   	   
   	    If Not IsDate(restore_time) Then
   			bfde4b54-0db7-4817-8032-87127bf19bb9 "Can't set f(x) view time to <" & restore_time & ">."
   		End If
   		
   		'---------------------------------------------------------
   		            
   	    ' go through the whole file, copy line by line, and replace the two archive variable names:
   	    While Not f2.eof
   			restore_entry=f2.lineinputstring
   			restore_entry= Replace(restore_entry, source_name1, target_name1)
   			restore_entry= Replace(restore_entry, source_name2, target_name2)
   			restore_entry= Replace(restore_entry, source_name3, target_name3)
   			restore_entry= Replace(restore_entry, source_name4, target_name4)
   			restore_entry= Replace(restore_entry, source_name5, target_name5)
   			restore_entry= Replace(restore_entry, source_name6, target_name6)
   			restore_entry= Replace(restore_entry, source_name7, target_name7)
   			restore_entry= Replace(restore_entry, source_name8, target_name8)
   			restore_entry= Replace(restore_entry, source_name9, target_name9)
   			f.lineprint(restore_entry)		
   		Wend
   		
   		f2.Close
   	    f.Close
   	       
   	    bb0abc73-aec8-40d0-9880-0280a6a3de42
   		Delay(2)
   		bec8f1e5-2ab1-45f6-ad91-1d37c469eb91 0502_Trend Historical, 0
   	            
   	    bfde4b54-0db7-4817-8032-87127bf19bb9 "Restored archive <" & archive_path & "> to <" & current_path &"> at " & restore_time & "."
   	    
   	    Set f2= Nothing
   	    Set f= Nothing
   		Else
   			
   		bb0abc73-aec8-40d0-9880-0280a6a3de42
   		bfde4b54-0db7-4817-8032-87127bf19bb9 "Long-term archive <" & archive_path & "> not found."
   	End If
   	
       Set fs= Nothing
       

VB script "LHmiView_vbsFECreateFolder"
   On Error Resume Next
   
   '-----------------------DEFINE PARAMETERS-------------------------------------------
   'kindOfOperatingSystem: 0 = Windows, 1 = Windows CE
   ' tempFs: Reference on temporary fileSystem Object
   ' fs: Reference on fileSystem Object
   ' f: Reference on file Object
   Dim kindOfOperatingSystem, tempFs, f, fs, file
   
   '--------------------Prove which Operating System is running------------------------
   'Set tempFs = CreateObject("Scripting.FileSystemObject")
   
   'If Err.Number = 0 Then
   '	kindOfOperatingSystem = 0 'Windows / PC based
   'Else
   	kindOfOperatingSystem = 1 'Windows CE / Panel based
   'End If
   
   Set tempFs= Nothing
   Err.Clear
   
   '-----------------create new folder-----------------------
   Dim newfolder
   
   If SmartTags("NewFolder") = "" Then 
     SmartTags("FEStatus") = "Folder name empty"
     Exit Sub
   End If
   
   newfolder = SmartTags("Folder") & SmartTags("NewFolder")
   
   'Windows CE / Panel based
   If kindOfOperatingSystem Then    
     Set fs = CreateObject("FileCtl.FileSystem")
     If fs.Dir(newfolder) = "" Then
       fs.MkDir(newfolder)
       If Err.Number = 0 Then
         SmartTags("FEStatus") = "Folder " & newfolder & " created"
       Else
         SmartTags("FEStatus") = "Could not create folder " & newfolder
       End If
     Else
       SmartTags("FEStatus") = "Folder exists already"
     End If
     
   ' Windows / PC based
   Else
     Set fs = CreateObject("Scripting.FileSystemObject")
     If fs.FolderExists(newfolder) = False Then
       fs.CreateFolder(newfolder)
       If Err.Number = 0 Then
         SmartTags("FEStatus") = "Folder " & newfolder & " created"
       Else
         SmartTags("FEStatus") = "Could not create folder " & newfolder
       End If
     Else
       SmartTags("FEStatus") = "Folder exists already"
     End If
   End If
   
   Set fs = Nothing
   
   LHmiView_vbsFEReadFilesOfFolder SmartTags("Folder")
   LHmiView_vbsFEWriteFilePropertiesToTags SmartTags("index")

VB script "LHmiView_vbsFEDelete"
   On Error Resume Next
   
   '-----------------------DEFINE PARAMETERS-------------------------------------------
   'kindOfOperatingSystem: 0 = Windows, 1 = Windows CE
   ' tempFs: Reference on temporary fileSystem Object
   ' fs: Reference on fileSystem Object
   ' f: Reference on file Object
   Dim kindOfOperatingSystem, tempFs, f, fs, file
   
   '--------------------Prove which Operating System is running------------------------
   'Set tempFs = CreateObject("Scripting.FileSystemObject")
   
   'If Err.Number = 0 Then
   '	kindOfOperatingSystem = 0 'Windows / PC based
   'Else
   	kindOfOperatingSystem = 1 'Windows CE / Panel based
   'End If
   
   Set tempFs= Nothing
   Err.Clear
   
   '-------------------------------Delete folder/file---------------------------------
   Dim i
   
   SmartTags("FEStatus") = "Deleting file..."
   i = SmartTags("fileChosen")
   
   ' Windows CE / Panel based
   If kindOfOperatingSystem Then    
     Set fs = CreateObject("FileCtl.FileSystem")
     Set f = CreateObject("FileCtl.File")
     If i > 0 And SmartTags("File_"&i) <> "" Then
       If SmartTags("isFolder_"&i) <> 0 Then
         fs.RmDir SmartTags("File_"&i)
         If Err.Number = 0 Then
           SmartTags("FEStatus") = "File / Folder deleted: " & SmartTags("File_"&i) 
           SmartTags("File_"&i) = ""
         Else
           SmartTags("FEStatus") = "Could not delete file / folder: " & SmartTags("File_"&i)
         End If
       Else
         fs.kill SmartTags("File_"&i)
         If Err.Number = 0 Then
           SmartTags("FEStatus") = "File / Folder deleted: " & SmartTags("File_"&i) 
         Else
           SmartTags("FEStatus") = "Could not delete file / folder: " & SmartTags("File_"&i)
         End If
         SmartTags("File_"&i) = ""
       End If
     Else
       SmartTags("FEStatus") = "Choose file / folder"
     End If
     
   ' Windows / PC based
   Else
     Set fs = CreateObject("Scripting.FileSystemObject")
      If i > 0 And SmartTags("File_"&i) <> "" Then
       If SmartTags("isFolder_"&i) <> "False" Then
         fs.DeleteFolder(SmartTags("File_"&i))
         If Err.Number = 0 Then
           SmartTags("FEStatus") = "File / folder deleted: " & SmartTags("File_"&i) 
           SmartTags("File_"&i) = ""
         Else
           SmartTags("FEStatus") = "Could not delete file / folder: " & SmartTags("File_"&i)
         End If
       Else
         fs.DeleteFile(SmartTags("File_"&i))
         If Err.Number = 0 Then
           SmartTags("FEStatus") = "Folder / folder deleted: " & SmartTags("File_"&i) 
         Else
           SmartTags("FEStatus") = "Could not delete file/ folder: " & SmartTags("File_"&i)
         End If
         SmartTags("File_"&i) = ""
       End If
     Else
       SmartTags("FEStatus") = "Choose file / folder"
     End If
   End If
   
   Set fs = Nothing
   Set f = Nothing
   
   LHmiView_vbsFEReadFilesOfFolder SmartTags("Folder")
   LHmiView_vbsFEWriteFilePropertiesToTags SmartTags("index")

VB script "LHmiView_vbsFEMove"
   On Error Resume Next
   
   '-----------------------DEFINE PARAMETERS-------------------------------------------
   'kindOfOperatingSystem: 0 = Windows, 1 = Windows CE
   ' tempFs: Reference on temporary fileSystem Object
   ' fs: Reference on fileSystem Object
   ' f: Reference on file Object
   Dim kindOfOperatingSystem, tempFs, f, fs, file
   
   '--------------------Prove which Operating System is running------------------------
   'Set tempFs = CreateObject("Scripting.FileSystemObject")
   
   'If Err.Number = 0 Then
   '	kindOfOperatingSystem = 0 'Windows / PC based
   'Else
   	kindOfOperatingSystem = 1 'Windows CE / Panel based
   'End If
   
   Set tempFs= Nothing
   Err.Clear
   
   '-------------------------------Move folder/file---------------------------------
   Dim  newpath, singleFile, data
   
   ' Windows CE / Panel based
   If kindOfOperatingSystem Then
     If sender = 1 Then 'button "copy" pressed
   	  If SmartTags("copyusb") = True Then
   		    If SmartTags("aIsFolder_"&SmartTags("AfileChosen")) = 0 Then
   		      SmartTags("bufferFile") = SmartTags("AFile_"&SmartTags("AfileChosen"))
   		      SmartTags("bufferFolder") = SmartTags("AFolder")
   		      SmartTags("bufferCopyCut") = True
   		      SmartTags("bufferIsFolder") = SmartTags("AisFolder_"&SmartTags("AfileChosen"))
   		      SmartTags("FEStatus") = "File " & SmartTags("bufferFile") & " copied"
   		    Else
   		      SmartTags("FEStatus") = "Cannot copy folder"
   			End If
   	  Else
   		   If SmartTags("IsFolder_"&SmartTags("fileChosen")) = 0 Then
   		      SmartTags("bufferFile") = SmartTags("File_"&SmartTags("fileChosen"))
   		      SmartTags("bufferFolder") = SmartTags("Folder")
   		      SmartTags("bufferCopyCut") = True
   		      SmartTags("bufferIsFolder") = SmartTags("isFolder_"&SmartTags("fileChosen"))
   		      SmartTags("FEStatus") = "File " & SmartTags("bufferFile") & " copied"
   		    Else
   		      SmartTags("FEStatus") = "Cannot copy folder"
   		   End If
   	  End If
   	  
     
     ElseIf sender = 3 Then 'button "cut" is pressed
   	  If SmartTags("copyusb") = True Then
   		    SmartTags("bufferFile") = SmartTags("AFile_"&SmartTags("AfileChosen"))
   		    SmartTags("bufferFolder") = SmartTags("AFolder")
   		    SmartTags("bufferCopyCut") = False 
   		    SmartTags("bufferIsFolder") = SmartTags("AisFolder_"&SmartTags("AfileChosen"))
   		    SmartTags("FEStatus") = "File " & SmartTags("bufferFile") & " cut"
   	  Else
   		  	SmartTags("bufferFile") = SmartTags("File_"&SmartTags("fileChosen"))
   		    SmartTags("bufferFolder") = SmartTags("Folder")
   		    SmartTags("bufferCopyCut") = False 
   		    SmartTags("bufferIsFolder") = SmartTags("isFolder_"&SmartTags("fileChosen"))
   		    SmartTags("FEStatus") = "File " & SmartTags("bufferFile") & " cut"   
   	  End If
   	  
   	  
     ElseIf sender = 2 Then 'button "move" pressed
       singleFile = Replace (SmartTags("bufferFile"),  SmartTags("bufferFolder"), "")
       newpath = SmartTags("Folder") & singleFile  
       If SmartTags("bufferCopyCut") = False Then   
         If SmartTags("bufferIsFolder") <> 0 Then
           Set fs = CreateObject("FileCtl.FileSystem")
           fs.MoveFile SmartTags("bufferFile"), newpath
         Else
           Set fs = CreateObject("FileCtl.FileSystem")
           fs.FileCopy SmartTags("bufferFile"), newpath
           fs.kill SmartTags("bufferFile")
         End If
       Else
         Set fs = CreateObject("FileCtl.FileSystem")
         fs.FileCopy SmartTags("bufferFile"), newpath
       End If 
       SmartTags("FEStatus") = "File " & SmartTags("bufferFile") & " pasted"
       LHmiView_vbsFEReadFilesOfFolder SmartTags("Folder")
       LHmiView_vbsFEWriteFilePropertiesToTags SmartTags("index")
     End If
   ' Windows / PC based
   Else
     If sender = 1 Then 'button "copy" pressed
   	  If SmartTags("copyusb") = True Then
   	    SmartTags("bufferFile") = SmartTags("aFile_"&SmartTags("AfileChosen"))
   	    SmartTags("bufferFolder") = SmartTags("AFolder")
   	    SmartTags("bufferCopyCut") = True
   	    SmartTags("bufferIsFolder") = SmartTags("aisFolder_"&SmartTags("AfileChosen"))
   	    SmartTags("FEStatus") = "File " & SmartTags("bufferFile") & " copied"
   	  Else
   		SmartTags("bufferFile") = SmartTags("File_"&SmartTags("fileChosen"))
   	    SmartTags("bufferFolder") = SmartTags("Folder")
   	    SmartTags("bufferCopyCut") = True
   	    SmartTags("bufferIsFolder") = SmartTags("isFolder_"&SmartTags("fileChosen"))
   	    SmartTags("FEStatus") = "File " & SmartTags("bufferFile") & " copied"
   	  End If
   	  
     
     ElseIf sender = 3 Then 'button "cut" is pressed
   	  If SmartTags("copyusb") = True Then
   		    SmartTags("bufferFile") = SmartTags("File_"&SmartTags("AfileChosen"))
   		    SmartTags("bufferFolder") = SmartTags("AFolder")
   		    SmartTags("bufferCopyCut") = False 
   		    SmartTags("bufferIsFolder") = SmartTags("aisFolder_"&SmartTags("AfileChosen"))
   		    SmartTags("FEStatus") = "File " & SmartTags("bufferFile") & " cut"
   	  Else
   		    SmartTags("bufferFile") = SmartTags("File_"&SmartTags("AfileChosen"))
   		    SmartTags("bufferFolder") = SmartTags("AFolder")
   		    SmartTags("bufferCopyCut") = False 
   		    SmartTags("bufferIsFolder") = SmartTags("aisFolder_"&SmartTags("AfileChosen"))
   		    SmartTags("FEStatus") = "File " & SmartTags("bufferFile") & " cut"
   	  End If    
   	  
     ElseIf sender = 2 Then 'button "move" pressed
       singleFile = Replace (SmartTags("bufferFile"),  SmartTags("bufferFolder"), "")
       newpath = SmartTags("Folder") & singleFile  
       Set fs = CreateObject("Scripting.FileSystemObject")
       If SmartTags("bufferCopyCut") = False Then
         If SmartTags("bufferIsFolder") = "True" Then
           data = fs.GetFolder(SmartTags("bufferFile"))
           fs.MoveFolder data, newpath
         Else
           data = fs.GetFile(SmartTags("bufferFile"))
           fs.MoveFile data, newpath
         End If
       Else
         If SmartTags("bufferIsFolder") = "True" Then
           data = fs.GetFolder(SmartTags("bufferFile"))
           fs.CopyFolder data, newpath
         Else
           data = fs.GetFile(SmartTags("bufferFile"))
           fs.CopyFile data, newpath
         End If
       End If
       If Err.Number <> 0 Then
         SmartTags("FEStatus") = Err.Description & "Could not paste file / folder"
       Else
         SmartTags("FEStatus") = "File / Folder " & SmartTags("bufferFile") & " pasted"
       End If
       LHmiView_vbsFEReadFilesOfFolder SmartTags("Folder")
       LHmiView_vbsFEWriteFilePropertiesToTags SmartTags("index")
     End If
   End If

VB script "LHmiView_vbsFEPreviousFolder"
   On Error Resume Next
   
   Dim folder, prevFolder
   
   If SmartTags("Search") = True Then
     SmartTags("Search") = False
     LHmiView_vbsFEReadFilesOfFolder(SmartTags("FEsearchFolder"))
     LHmiView_vbsFEWriteFilePropertiesToTags 1
   Else
   	If Len(SmartTags("Folder")) > 1 Then
   	    folder = Left (SmartTags("Folder"),  InStrRev (SmartTags("Folder"), "\")-1)
   	    prevFolder = Left (folder, InStrRev (folder, "\"))
   	    LHmiView_vbsFEReadFilesOfFolder(prevFolder)
   	    LHmiView_vbsFEWriteFilePropertiesToTags 1
   	    SmartTags("index") = 1
   	    SmartTags("FEStatus") = "Folder " & prevFolder & " opened"
   	Else
   	    SmartTags("FEStatus") = "Operation not possible"
   	End If
   End If

VB script "LHmiView_vbsFEReadFilesOfFolder"
   On Error Resume Next
   
   '-----------------------DEFINE PARAMETERS-------------------------------------------
   'kindOfOperatingSystem: 0 = Windows, 1 = Windows CE
   ' tempFs: Reference on temporary fileSystem Object
   ' fs: Reference on fileSystem Object
   ' f: Reference on file Object
   Dim kindOfOperatingSystem, tempFs, f, fs, file
   
   '--------------------Prove which Operating System is running------------------------
   'Set tempFs = CreateObject("Scripting.FileSystemObject")
   
   'If Err.Number = 0 Then
   '	kindOfOperatingSystem = 0 'Windows / PC based
   'Else
   	kindOfOperatingSystem = 1 'Windows CE / Panel based
   'End If
   
   Set tempFs= Nothing
   Err.Clear
   
   '-------------------------------Read files of folder---------------------------------
   Dim isFolder, counter, index, textStream, folder, dataInFolder, fileList
   
   index = 1
   
   ' Windows CE / Panel based
   If kindOfOperatingSystem Then 
     If folderpar = "" Then
       folderpar = "\"
     End If
        
     Set fs = CreateObject("FileCtl.FileSystem")
     Set f = CreateObject("FileCtl.File")
     If fs.Dir("\flash\106226404_Tools") = "" Then   fs.MkDir("\flash\106226404_Tools")
     f.open "\flash\106226404_Tools\LHmiView_FileList.txt", 2 'textfile where the files are stored
     
     file = fs.dir(folderpar & "*")
     counter = 0
     index = 1
     f.lineprint(folderpar)
     f.lineprint("-1")
     f.LinePrint "#106226404_FE_Site_"&index
     
     Do While file <> "" 
       If (counter < 10) Then  'write 10 files (pathname and isFolder) to textfile
         If ((fs.GetAttr(folderpar & file) And 16) <> 0 ) Then
           isFolder = True
         Else
           isFolder = False
         End If
         f.LinePrint(folderpar & file)
         f.LinePrint(isFolder)
         file = fs.dir
         counter = counter + 1
       Else
         counter = 0
         index = index + 1
         f.LinePrint "#106226404_FE_Site_"&index 
       End If
     Loop
     
     f.Close
     
   ' Windows / PC based
   Else
     If (folderpar = "") Then
       folderpar = "C:\"
     End If
     
     Set fs = CreateObject("Scripting.FileSystemObject")
     fileList = "C:\106226404_Tools\LHmiView_FileList.txt"
     If Not fs.FolderExists("C:\106226404_Tools") Then fs.CreateFolder "C:\106226404_Tools"
     If Not fs.FileExists(fileList) Then fs.CreateTextFile fileList
     Set f = fs.GetFile(fileList)
     Set textStream = f.OpenAsTextStream(2,-2)
     
     counter = 0
     index = 1
     textStream.WriteLine(folderpar)
     textStream.WriteLine("-1")
     textStream.WriteLine "#106226404_FE_Site_"&index
     
     Set folder = fs.GetFolder(folderpar)
     
     Set dataInFolder = folder.SubFolders
     For Each file In dataInFolder
       If Not file.Attributes And 2 Then
         If (counter < 10) Then 'write 10 files (pathname and isFolder) to textfile
           textStream.WriteLine(file.Path)
           textStream.WriteLine("True")
           counter = counter + 1
         Else
           counter = 0
           index = index + 1
           textStream.WriteLine "#106226404_FE_Site_"&index 
         End If
       End If
     Next
     
     Set dataInFolder = folder.Files
     For Each file In dataInFolder
       If Not file.Attributes And 2 Then
         If (counter < 10) Then 'write 10 folder (pathname and isFolder) to textfile
           textStream.WriteLine(file.Path)
           textStream.WriteLine("False")
           counter = counter + 1
         Else
           counter = 0
           index = index + 1
           textStream.WriteLine "#106226404_FE_Site_"&index 
         End If
       End If
     Next
   
     textStream.Close
     Set folder = Nothing
     Set dataInFolder = Nothing
     Set textStream = Nothing
   
   End If
   Set fs = Nothing
   Set f = Nothing

VB script "LHmiView_vbsFERename"
   On Error Resume Next
   
   '-----------------------DEFINE PARAMETERS-------------------------------------------
   'kindOfOperatingSystem: 0 = Windows, 1 = Windows CE
   ' tempFs: Reference on temporary fileSystem Object
   ' fs: Reference on fileSystem Object
   ' f: Reference on file Object
   Dim kindOfOperatingSystem, tempFs, f, fs,file
   
   '--------------------Prove which Operating System is running------------------------
   'Set tempFs = CreateObject("Scripting.FileSystemObject")
   
   'If Err.Number = 0 Then
   '	kindOfOperatingSystem = 0 'Windows / PC based
   'Else
   	kindOfOperatingSystem = 1 'Windows CE / Panel based
   'End If
   
   Set tempFs= Nothing
   Err.Clear
   
   '-------------------------------Rename folder/file---------------------------------
   Dim i, newName, ext, fileName, folder
   
   i = SmartTags("fileChosen")
   fileName = SmartTags("File_"&i)
   
   If fileName <> "" And SmartTags("NewName") <> "" Then
     
     ' Windows CE / Panel based
     If kindOfOperatingSystem Then    
       Set fs = CreateObject("FileCtl.FileSystem")
       If SmartTags("IsFolder_"&i) <> 0 Then 'Rename folder
         newName = SmartTags("Folder") & SmartTags("NewName")
         fs.MoveFile fileName, newName
         If Err.Number = 0 Then
           SmartTags("FEStatus") = "Folder renamed in: " & newName
         Else
           SmartTags("FEStatus") = "Could not rename folder: " & fileName
         End If
       Else 'Keep file extension
         ext = Right(fileName, Len(fileName)-InStrRev(fileName, "."))
         newName = SmartTags("Folder") & SmartTags("NewName") & "." & ext
         fs.MoveFile fileName, newName
         If Err.Number = 0 Then
           SmartTags("FEStatus") = "File renamed in: " & newName
         Else
           SmartTags("FEStatus") = "Could not rename file:" & fileName
         End If    
       End If
       
     ' Windows / PC based
     Else
       Set fs = CreateObject("Scripting.FileSystemObject")
       If SmartTags("IsFolder_"&i) <> "False" Then 'Rename folder
         Set folder = fs.GetFolder(fileName)
         newName = SmartTags("Folder") & SmartTags("NewName")
         fs.MoveFolder fileName, newName
         If Err.Number = 0 Then
           SmartTags("FEStatus") = "Folder renamed in: " & newName
         Else
           SmartTags("FEStatus") = "Error :" & Err.Description & " Could not rename folder: " & fileName
         End If
         Set folder = Nothing
       Else 'Keep file extension
        Set file = fs.GetFile(fileName)
         ext = Right(fileName, Len(fileName)-InStrRev(fileName, "."))
         newName = SmartTags("NewName") & "." & ext
         file.Name = newName
         If Err.Number = 0 Then
           SmartTags("FEStatus") = "File renamed in: " & newName
         Else
           SmartTags("FEStatus") = "Could not rename file: " & fileName
         End If    
         Set file = Nothing
       End If 
     End If
     Set fs = Nothing
    
   Else
     SmartTags("FEStatus") = "No file / folder chosen or name empty"
   End If
   Set fs = Nothing
   LHmiView_vbsFEReadFilesOfFolder SmartTags("Folder")
   LHmiView_vbsFEWriteFilePropertiesToTags SmartTags("index")
     

VB script "LHmiView_vbsFESearch"
   On Error Resume Next
   
   '-----------------------DEFINE PARAMETERS-------------------------------------------
   'kindOfOperatingSystem: 0 = Windows, 1 = Windows CE
   ' tempFs: Reference on temporary fileSystem Object
   ' fs: Reference on fileSystem Object
   ' f: Reference on file Object
   Dim kindOfOperatingSystem, tempFs, f, fs, file
   
   '--------------------Prove which Operating System is running------------------------
   'Set tempFs = CreateObject("Scripting.FileSystemObject")
   
   'If Err.Number = 0 Then
   '	kindOfOperatingSystem = 0 'Windows / PC based
   'Else
   	kindOfOperatingSystem = 1 'Windows CE / Panel based
   'End If
   
   Set tempFs= Nothing
   Err.Clear
   
   '-------------------------------Search folder/file---------------------------------
   Dim i, j, index, line, buffer(), searchString
   
   If SmartTags("FEsearchString") <> "" Then
     SmartTags("FEStatus") = "Searching for text: " & SmartTags("FEsearchString") & "..."
     
     'Windows CE / Panel based
     If kindOfOperatingSystem Then
       Set f = CreateObject("filectl.file")
       Set fs = CreateObject("filectl.Filesystem")
       file = "\flash\106226404_Tools\LHmiView_FileList.txt"
       f.open file, 1 
       i=1
       j=1
       searchString = LCase(SmartTags("FEsearchString")) 
       Do While f.EOF = False 'Check number of lines for Array Definition
         f.LineInputString
         i=i+1
       Loop
       ReDim buffer(i)
       'Reinitialize
       i=1
       f.close
       f.open file,1
       Do While f.EOF = False
         line = LCase(f.LineInputString)
          If InStr(1,line,searchString,0) <> 0 Then
            buffer(i) = line
            buffer(i+1) = f.LineInputString
            i = i+2
            bfde4b54-0db7-4817-8032-87127bf19bb9("Found: "&line)
          End If
       Loop
       f.Close
       If i>1 Then
         SmartTags("FEsearchFolder") = SmartTags("Folder")
         f.open "\flash\106226404_Tools\LHmiView_SearchList.txt", 2  
         index = 1
         f.LinePrint SmartTags("Folder")
         f.LinePrint "#106226404_FE_Site_"&index
         For j=1 To i
           f.LinePrint(buffer(j))
           bfde4b54-0db7-4817-8032-87127bf19bb9("Written: " &buffer(j))
           If (j Mod 20) = 0 Then
             index = index+1
             f.LinePrint "#106226404_FE_Site_"&index
           End If
         Next
         f.close
         fs.kill "\flash\106226404_Tools\LHmiView_FileList.txt"
         fs.FileCopy "\flash\106226404_Tools\LHmiView_SearchList.txt", "\flash\106226404_Tools\LHmiView_FileList.txt"
         fs.kill "\flash\106226404_Tools\LHmiView_SearchList.txt"
         LHmiView_vbsFEWriteFilePropertiesToTags 1
       End If
       SmartTags("FEStatus") = (i-1)/2 & " Files found with text: " & SmartTags("FEsearchString") 
       Set f = Nothing
       Set fs = Nothing
       
     'Windows / PC based
     Else
       Set fs = CreateObject("Scripting.FileSystemObject")
       file = "C:\106226404_Tools\LHmiView_FileList.txt"
       Set f = fs.OpenTextFile (file, 1) 
       i=1
       j=1
       searchString = LCase(SmartTags("FEsearchString")) 
       Do While f.AtEndOfStream <> True 'Check number of lines for Array Definition
         f.ReadLine
         i=i+1
       Loop
       ReDim buffer(i)
       'Reinitialize
       i=1
       f.Close
       Set f = fs.OpenTextFile (file, 1)
       Do While f.AtEndOfStream <> True
         line = LCase(f.ReadLine)
         If InStr(1,line,searchString,0) <> 0 Then
           buffer(i) = line
           buffer(i+1) = f.ReadLine
           i = i+2
         End If
       Loop
       f.Close
       If i>1 Then
         SmartTags("FEsearchFolder") = SmartTags("Folder")
         file = "C:\106226404_Tools\LHmiView_SearchList.txt"
         If Not fs.FileExists(file) Then fs.CreateTextFile file
         Set f = fs.OpenTextFile (file, 2)
         index = 1
         f.WriteLine SmartTags("Folder")
         f.WriteLine "#106226404_FE_Site_"&index
         For j=1 To i
           f.WriteLine(buffer(j))
           bfde4b54-0db7-4817-8032-87127bf19bb9("Written: " &buffer(j))
           If (j Mod 20) = 0 Then
             index = index+1
             f.WriteLine "#106226404_FE_Site_"&index
           End If
         Next
         f.Close
         fs.DeleteFile "C:\106226404_Tools\LHmiView_FileList.txt"
         fs.CopyFile "C:\106226404_Tools\LHmiView_SearchList.txt", "C:\106226404_Tools\LHmiView_FileList.txt"
         fs.DeleteFile "C:\106226404_Tools\LHmiView_SearchList.txt"
         LHmiView_vbsFEWriteFilePropertiesToTags 1
       End If
       SmartTags("FEStatus") = (i-1)/2 & " Files found with text: " & SmartTags("FEsearchString") 
       Set f = Nothing
       Set fs = Nothing          
     End If        
   Else
     SmartTags("FEStatus") = "Search text empty"
   End If      

VB script "LHmiView_vbsFEShowFiles"
   On Error Resume Next
   
   '-----------------------DEFINE PARAMETERS-------------------------------------------
   'kindOfOperatingSystem: 0 = Windows, 1 = Windows CE
   ' tempFs: Reference on temporary fileSystem Object
   ' fs: Reference on fileSystem Object
   ' f: Reference on file Object
   Dim kindOfOperatingSystem, tempFs, f, fs, file
   
   '--------------------Prove which Operating System is running------------------------
   'Set tempFs = CreateObject("Scripting.FileSystemObject")
   
   'If Err.Number = 0 Then
   '	kindOfOperatingSystem = 0 'Windows / PC based
   'Else
   	kindOfOperatingSystem = 1 'Windows CE / Panel based
   'End If
   
   Set tempFs= Nothing
   Err.Clear
   
   '-----------------show files -----------------------
   Dim fileName, ext, obj
   'Windows CE / Panel based
   
   If kindOfOperatingSystem Then  
     If SmartTags("File_"&SmartTags("fileChosen")) <> "" Then
       If SmartTags("IsFolder_"&SmartTags("fileChosen")) <> 0 Then
           LHmiView_vbsFEReadFilesOfFolder(SmartTags("File_"&SmartTags("fileChosen"))&"\")
           LHmiView_vbsFEWriteFilePropertiesToTags 1
           SmartTags("index") = 1
       Else
         fileName = SmartTags("File_"&SmartTags("fileChosen")) 
         ext = LCase(Right(fileName, Len(fileName)-InStrRev(fileName, "."))) 
         fileName = Chr(34) & fileName & Chr(34) ' Add " for spaces in fileName
       ' ExcelViewer: *.xlsx, *.xls, *.xlt
       ' WordViewer: *.docx, *.rtf, *.doc
       ' PdfViewer *.pdf
       ' Internet Explorer *.html
       ' Mediaplayer *.mpa, *.mp2, *.mp3, *.wma, *wav, *.mpg, *.mpeg, *.mpe, *.asf, *.wmv, *.avi
         If ext = "xlsx" Or ext = "xls" Or ext = "xlt" Or _
         ext = "docx" Or ext = "rtf" Or ext = "doc" Or _
         ext = "pdf" Or _
         ext = "html" Or _
         ext = "mpa" Or ext = "mp2" Or ext = "mp3" Or ext = "wma" Or ext = "wav" Or ext = "mpg" Or ext = "mpeg" Or ext = "mpe" Or ext = "asf" Or ext = "wmv" Or ext = "avi" Then
             bf5b406f-e168-4434-a306-9566226aa38b fileName, "", $3$hmiShowNormal$, $3$hmiNo$
         Else
           SmartTags("FEStatus") = "Cannot open file"
         End If  
       End If
     End If
   'Windows / PC based 
   Else
     If SmartTags("File_"&SmartTags("fileChosen")) <> "" Then
       If SmartTags("IsFolder_"&SmartTags("fileChosen")) <> "False" Then
         LHmiView_vbsFEReadFilesOfFolder(SmartTags("File_"&SmartTags("fileChosen"))&"\")
         LHmiView_vbsFEWriteFilePropertiesToTags 1
         SmartTags("index") = 1
       Else  
         fileName = SmartTags("File_"&SmartTags("fileChosen")) 
         Set obj = CreateObject("Wscript.Shell")
         obj.Run fileName
       End If
     Else
       SmartTags("FEStatus") = "No file or folder chosen"
     End If
   End If

VB script "LHmiView_vbsFEWriteFilePropertiesToTags"
   On Error Resume Next
   
   '-----------------------DEFINE PARAMETERS-------------------------------------------
   'kindOfOperatingSystem: 0 = Windows, 1 = Windows CE
   ' tempFs: Reference on temporary fileSystem Object
   ' fs: Reference on fileSystem Object
   ' f: Reference on file Object
   Dim kindOfOperatingSystem, tempFs, f, fs, file
   
   '--------------------Prove which Operating System is running------------------------
   'Set tempFs = CreateObject("Scripting.FileSystemObject")
   
   'If Err.Number = 0 Then
   '	kindOfOperatingSystem = 0 'Windows / PC based
   'Else
   	kindOfOperatingSystem = 1 'Windows CE / Panel based
   'End If
   
   Set tempFs= Nothing
   Err.Clear
   
   '-----------------create new folder-----------------------
   Dim i
   
   If kindOfOperatingSystem Then    
     Set fs = CreateObject("FileCtl.FileSystem")
     Set f = CreateObject("FileCtl.File")
     file = "\flash\106226404_Tools\LHmiView_FileList.txt"
     SmartTags("NextPossible") = True
     If fs.Dir(file) <> "" Then
       f.open file, 1
       SmartTags("Folder") = f.LineInputString
       Do While f.LineInputString <>  "#106226404_FE_Site_"&index  'find current position in file 
       Loop
       
       For i=1 To 10
         If f.EOF = False Then       
           SmartTags("File_" &i) = f.LineInputString
         Else  ' fill tags at the end of the file
           SmartTags("File_" &i) = ""
         End If
         If f.EOF = False Then
           SmartTags("isFolder_" &i) = f.LineInputString
         Else  
           SmartTags("isFolder_" &i) = ""     
         End If
       Next
       
       If f.EOF = True Then
         SmartTags("NextPossible") = False
       Else 
         SmartTags("NextPossible") = True
       End If
       f.Close 
       f.Close
     End If
   ' Windows / PC based
   Else
     Set fs = CreateObject("Scripting.FileSystemObject")
     file = "C:\106226404_Tools\LHmiView_FileList.txt"
     If Not fs.FileExists(file) Then Exit Sub
     Set f = fs.OpenTextFile (file, 1)
     SmartTags("Folder") = f.ReadLine
     Do While f.ReadLine <>  "#106226404_FE_Site_"&index  'find current position in file 
     Loop
     
     For i=1 To 10
       If f.AtEndOfStream = False Then       
         SmartTags("File_" &i) = f.ReadLine
       Else  ' fill tags at the end of the file
         SmartTags("File_" &i) = ""
       End If
       If f.AtEndOfStream = False Then
         SmartTags("isFolder_" &i) = f.ReadLine
       Else  
         SmartTags("isFolder_" &i) = ""     
       End If
     Next
     
     If f.AtEndOfStream = True Then
       SmartTags("NextPossible") = False
     Else 
       SmartTags("NextPossible") = True
     End If
     f.Close    
   End If
   Set fs = Nothing
   Set f = Nothing

VB script "LHmiView_vbsFESearch_1"
   On Error Resume Next
   
   '-----------------------DEFINE PARAMETERS-------------------------------------------
   'kindOfOperatingSystem: 0 = Windows, 1 = Windows CE
   ' tempFs: Reference on temporary fileSystem Object
   ' fs: Reference on fileSystem Object
   ' f: Reference on file Object
   Dim kindOfOperatingSystem, tempFs, f, fs, file
   
   '--------------------Prove which Operating System is running------------------------
   'Set tempFs = CreateObject("Scripting.FileSystemObject")
   
   'If Err.Number = 0 Then
   '	kindOfOperatingSystem = 0 'Windows / PC based
   'Else
   	kindOfOperatingSystem = 1 'Windows CE / Panel based
   'End If
   
   Set tempFs= Nothing
   Err.Clear
   
   '-------------------------------Search folder/file---------------------------------
   Dim i, j, index, line, buffer(), searchString
   
   If SmartTags("AFEsearchString") <> "" Then
     SmartTags("AFEStatus") = "Searching for text: " & SmartTags("AFEsearchString") & "..."
     
     'Windows CE / Panel based
     If kindOfOperatingSystem Then
       Set f = CreateObject("filectl.file")
       Set fs = CreateObject("filectl.Filesystem")
       file = "\flash\106226404_Tools\LHmiView_FileListB.txt"
       f.open file, 1 
       i=1
       j=1
       searchString = LCase(SmartTags("AFEsearchString")) 
       Do While f.EOF = False 'Check number of lines for Array Definition
         f.LineInputString
         i=i+1
       Loop
       ReDim buffer(i)
       'Reinitialize
       i=1
       f.close
       f.open file,1
       Do While f.EOF = False
         line = LCase(f.LineInputString)
          If InStr(1,line,searchString,0) <> 0 Then
            buffer(i) = line
            buffer(i+1) = f.LineInputString
            i = i+2
            bfde4b54-0db7-4817-8032-87127bf19bb9("Found: "&line)
          End If
       Loop
       f.Close
       If i>1 Then
         SmartTags("AFEsearchFolder") = SmartTags("AFolder")
         f.open "\flash\106226404_Tools\LHmiView_SearchListB.txt", 2  
         index = 1
         f.LinePrint SmartTags("AFolder")
         f.LinePrint "#106226404_FE_Site_"&index
         For j=1 To i
           f.LinePrint(buffer(j))
           bfde4b54-0db7-4817-8032-87127bf19bb9("Written: " &buffer(j))
           If (j Mod 20) = 0 Then
             index = index+1
             f.LinePrint "#106226404_FE_Site_"&index
           End If
         Next
         f.close
         fs.kill "\flash\106226404_Tools\LHmiView_FileListB.txt"
         fs.FileCopy "\flash\106226404_Tools\LHmiView_SearchListB.txt", "\flash\106226404_Tools\LHmiView_FileListB.txt"
         fs.kill "\flash\106226404_Tools\LHmiView_SearchListB.txt"
         LHmiView_vbsFEWriteFilePropertiesToTags_1 1
       End If
       SmartTags("AFEStatus") = (i-1)/2 & " Files found with text: " & SmartTags("AFEsearchString") 
       Set f = Nothing
       Set fs = Nothing
       
     'Windows / PC based
     Else
       Set fs = CreateObject("Scripting.FileSystemObject")
       file = "C:\106226404_Tools\LHmiView_FileListB.txt"
       Set f = fs.OpenTextFile (file, 1) 
       i=1
       j=1
       searchString = LCase(SmartTags("AFEsearchString")) 
       Do While f.AtEndOfStream <> True 'Check number of lines for Array Definition
         f.ReadLine
         i=i+1
       Loop
       ReDim buffer(i)
       'Reinitialize
       i=1
       f.Close
       Set f = fs.OpenTextFile (file, 1)
       Do While f.AtEndOfStream <> True
         line = LCase(f.ReadLine)
         If InStr(1,line,searchString,0) <> 0 Then
           buffer(i) = line
           buffer(i+1) = f.ReadLine
           i = i+2
         End If
       Loop
       f.Close
       If i>1 Then
         SmartTags("AFEsearchFolder") = SmartTags("AFolder")
         file = "C:\106226404_Tools\LHmiView_SearchListB.txt"
         If Not fs.FileExists(file) Then fs.CreateTextFile file
         Set f = fs.OpenTextFile (file, 2)
         index = 1
         f.WriteLine SmartTags("AFolder")
         f.WriteLine "#106226404_FE_Site_"&index
         For j=1 To i
           f.WriteLine(buffer(j))
           bfde4b54-0db7-4817-8032-87127bf19bb9("Written: " &buffer(j))
           If (j Mod 20) = 0 Then
             index = index+1
             f.WriteLine "#106226404_FE_Site_"&index
           End If
         Next
         f.Close
         fs.DeleteFile "C:\106226404_Tools\LHmiView_FileListB.txt"
         fs.CopyFile "C:\106226404_Tools\LHmiView_SearchListB.txt", "C:\106226404_Tools\LHmiView_FileListB.txt"
         fs.DeleteFile "C:\106226404_Tools\LHmiView_SearchListB.txt"
         LHmiView_vbsFEWriteFilePropertiesToTags_1 1
       End If
       SmartTags("AFEStatus") = (i-1)/2 & " Files found with text: " & SmartTags("AFEsearchString") 
       Set f = Nothing
       Set fs = Nothing          
     End If        
   Else
     SmartTags("AFEStatus") = "Search text empty"
   End If      

VB script "LHmiView_vbsFEWriteFilePropertiesToTags_1"
   On Error Resume Next
   
   '-----------------------DEFINE PARAMETERS-------------------------------------------
   'kindOfOperatingSystem: 0 = Windows, 1 = Windows CE
   ' tempFs: Reference on temporary fileSystem Object
   ' fs: Reference on fileSystem Object
   ' f: Reference on file Object
   Dim kindOfOperatingSystem, tempFs, f, fs, file
   
   '--------------------Prove which Operating System is running------------------------
   'Set tempFs = CreateObject("Scripting.FileSystemObject")
   
   'If Err.Number = 0 Then
   '	kindOfOperatingSystem = 0 'Windows / PC based
   'Else
   	kindOfOperatingSystem = 1 'Windows CE / Panel based
   'End If
   
   Set tempFs= Nothing
   Err.Clear
   
   '-----------------create new folder-----------------------
   Dim i
   
   If kindOfOperatingSystem Then    
     Set fs = CreateObject("FileCtl.FileSystem")
     Set f = CreateObject("FileCtl.File")
     file = "\flash\106226404_Tools\LHmiView_FileListB.txt"
     SmartTags("ANextPossible") = True
     If fs.Dir(file) <> "" Then
       f.open file, 1
       SmartTags("AFolder") = f.LineInputString
       Do While f.LineInputString <>  "#106226404_FE_Site_"&index  'find current position in file 
       Loop
       
       For i=1 To 10
         If f.EOF = False Then       
           SmartTags("AFile_" &i) = f.LineInputString
         Else  ' fill tags at the end of the file
           SmartTags("AFile_" &i) = ""
         End If
         If f.EOF = False Then
           SmartTags("AisFolder_" &i) = f.LineInputString
         Else  
           SmartTags("AisFolder_" &i) = ""     
         End If
       Next
       
       If f.EOF = True Then
         SmartTags("ANextPossible") = False
       Else 
         SmartTags("ANextPossible") = True
       End If
       f.Close 
       f.Close
     End If
   ' Windows / PC based
   Else
     Set fs = CreateObject("Scripting.FileSystemObject")
     file = "C:\106226404_Tools\LHmiView_FileListB.txt"
     If Not fs.FileExists(file) Then Exit Sub
     Set f = fs.OpenTextFile (file, 1)
     SmartTags("AFolder") = f.ReadLine
     Do While f.ReadLine <>  "#106226404_FE_Site_"&index  'find current position in file 
     Loop
     
     For i=1 To 10
       If f.AtEndOfStream = False Then       
         SmartTags("aFile_" &i) = f.ReadLine
       Else  ' fill tags at the end of the file
         SmartTags("aFile_" &i) = ""
       End If
       If f.AtEndOfStream = False Then
         SmartTags("aisFolder_" &i) = f.ReadLine
       Else  
         SmartTags("aisFolder_" &i) = ""     
       End If
     Next
     
     If f.AtEndOfStream = True Then
       SmartTags("ANextPossible") = False
     Else 
       SmartTags("ANextPossible") = True
     End If
     f.Close    
   End If
   Set fs = Nothing
   Set f = Nothing

VB script "LHmiView_vbsFEPreviousFolder_1"
   On Error Resume Next
   
   Dim folder, prevFolder
   
   If SmartTags("ASearch") = True Then
     SmartTags("ASearch") = False
     LHmiView_vbsFEReadFilesOfFolder_1(SmartTags("AFEsearchFolder"))
     LHmiView_vbsFEWriteFilePropertiesToTags_1 1
   Else
   	If Len(SmartTags("AFolder")) > 1 Then
   	    folder = Left (SmartTags("AFolder"),  InStrRev (SmartTags("AFolder"), "\")-1)
   	    prevFolder = Left (folder, InStrRev (folder, "\"))
   	    LHmiView_vbsFEReadFilesOfFolder_1(prevFolder)
   	    LHmiView_vbsFEWriteFilePropertiesToTags_1 1
   	    SmartTags("Aindex") = 1
   	    SmartTags("AFEStatus") = "Folder " & prevFolder & " opened"
   	Else
   	    SmartTags("AFEStatus") = "Operation not possible"
   	End If
   End If

VB script "LHmiView_vbsFEReadFilesOfFolder_1"
   On Error Resume Next
   
   '-----------------------DEFINE PARAMETERS-------------------------------------------
   'kindOfOperatingSystem: 0 = Windows, 1 = Windows CE
   ' tempFs: Reference on temporary fileSystem Object
   ' fs: Reference on fileSystem Object
   ' f: Reference on file Object
   Dim kindOfOperatingSystem, tempFs, f, fs, file
   
   '--------------------Prove which Operating System is running------------------------
   'Set tempFs = CreateObject("Scripting.FileSystemObject")
   
   'If Err.Number = 0 Then
   '	kindOfOperatingSystem = 0 'Windows / PC based
   'Else
   	kindOfOperatingSystem = 1 'Windows CE / Panel based
   'End If
   
   Set tempFs= Nothing
   Err.Clear
   
   '-------------------------------Read files of folder---------------------------------
   Dim isFolder, counter, index, textStream, folder, dataInFolder, fileList
   
   index = 1
   
   ' Windows CE / Panel based
   If kindOfOperatingSystem Then 
     If folderpar = "" Then
       folderpar = "\"
     End If
        
     Set fs = CreateObject("FileCtl.FileSystem")
     Set f = CreateObject("FileCtl.File")
     If fs.Dir("\flash\106226404_Tools") = "" Then   fs.MkDir("\flash\106226404_Tools")
     f.open "\flash\106226404_Tools\LHmiView_FileListB.txt", 2 'textfile where the files are stored
     
     file = fs.dir(folderpar & "*")
     counter = 0
     index = 1
     f.lineprint(folderpar)
     f.lineprint("-1")
     f.LinePrint "#106226404_FE_Site_"&index
     
     Do While file <> "" 
       If (counter < 10) Then  'write 10 files (pathname and isFolder) to textfile
         If ((fs.GetAttr(folderpar & file) And 16) <> 0 ) Then
           isFolder = True
         Else
           isFolder = False
         End If
         f.LinePrint(folderpar & file)
         f.LinePrint(isFolder)
         file = fs.dir
         counter = counter + 1
       Else
         counter = 0
         index = index + 1
         f.LinePrint "#106226404_FE_Site_"&index 
       End If
     Loop
     
     f.Close
     
   ' Windows / PC based
   Else
     If (folderpar = "") Then
       folderpar = "C:\"
     End If
     
     Set fs = CreateObject("Scripting.FileSystemObject")
     fileList = "C:\106226404_Tools\LHmiView_FileListB.txt"
     If Not fs.FolderExists("C:\106226404_Tools") Then fs.CreateFolder "C:\106226404_Tools"
     If Not fs.FileExists(fileList) Then fs.CreateTextFile fileList
     Set f = fs.GetFile(fileList)
     Set textStream = f.OpenAsTextStream(2,-2)
     
     counter = 0
     index = 1
     textStream.WriteLine(folderpar)
     textStream.WriteLine("-1")
     textStream.WriteLine "#106226404_FE_Site_"&index
     
     Set folder = fs.GetFolder(folderpar)
     
     Set dataInFolder = folder.SubFolders
     For Each file In dataInFolder
       If Not file.Attributes And 2 Then
         If (counter < 10) Then 'write 10 files (pathname and isFolder) to textfile
           textStream.WriteLine(file.Path)
           textStream.WriteLine("True")
           counter = counter + 1
         Else
           counter = 0
           index = index + 1
           textStream.WriteLine "#106226404_FE_Site_"&index 
         End If
       End If
     Next
     
     Set dataInFolder = folder.Files
     For Each file In dataInFolder
       If Not file.Attributes And 2 Then
         If (counter < 10) Then 'write 10 folder (pathname and isFolder) to textfile
           textStream.WriteLine(file.Path)
           textStream.WriteLine("False")
           counter = counter + 1
         Else
           counter = 0
           index = index + 1
           textStream.WriteLine "#106226404_FE_Site_"&index 
         End If
       End If
     Next
   
     textStream.Close
     Set folder = Nothing
     Set dataInFolder = Nothing
     Set textStream = Nothing
   
   End If
   Set fs = Nothing
   Set f = Nothing

VB script "LHmiView_vbsFEShowFiles_1"
   On Error Resume Next
   
   '-----------------------DEFINE PARAMETERS-------------------------------------------
   'kindOfOperatingSystem: 0 = Windows, 1 = Windows CE
   ' tempFs: Reference on temporary fileSystem Object
   ' fs: Reference on fileSystem Object
   ' f: Reference on file Object
   Dim kindOfOperatingSystem, tempFs, f, fs, file
   
   '--------------------Prove which Operating System is running------------------------
   'Set tempFs = CreateObject("Scripting.FileSystemObject")
   
   'If Err.Number = 0 Then
   '	kindOfOperatingSystem = 0 'Windows / PC based
   'Else
   	kindOfOperatingSystem = 1 'Windows CE / Panel based
   'End If
   
   Set tempFs= Nothing
   Err.Clear
   
   '-----------------show files -----------------------
   Dim fileName, ext, obj
   'Windows CE / Panel based
   
   If kindOfOperatingSystem Then  
     If SmartTags("AFile_"&SmartTags("AfileChosen")) <> "" Then
       If SmartTags("AIsFolder_"&SmartTags("AfileChosen")) <> 0 Then
           LHmiView_vbsFEReadFilesOfFolder_1(SmartTags("AFile_"&SmartTags("AfileChosen"))&"\")
           LHmiView_vbsFEWriteFilePropertiesToTags_1 1
           SmartTags("Aindex") = 1
       Else
         fileName = SmartTags("AFile_"&SmartTags("AfileChosen")) 
         ext = LCase(Right(fileName, Len(fileName)-InStrRev(fileName, "."))) 
         fileName = Chr(34) & fileName & Chr(34) ' Add " for spaces in fileName
       ' ExcelViewer: *.xlsx, *.xls, *.xlt
       ' WordViewer: *.docx, *.rtf, *.doc
       ' PdfViewer *.pdf
       ' Internet Explorer *.html
       ' Mediaplayer *.mpa, *.mp2, *.mp3, *.wma, *wav, *.mpg, *.mpeg, *.mpe, *.asf, *.wmv, *.avi
         If ext = "xlsx" Or ext = "xls" Or ext = "xlt" Or _
         ext = "docx" Or ext = "rtf" Or ext = "doc" Or _
         ext = "pdf" Or _
         ext = "html" Or _
         ext = "mpa" Or ext = "mp2" Or ext = "mp3" Or ext = "wma" Or ext = "wav" Or ext = "mpg" Or ext = "mpeg" Or ext = "mpe" Or ext = "asf" Or ext = "wmv" Or ext = "avi" Then
             bf5b406f-e168-4434-a306-9566226aa38b fileName, "", $3$hmiShowNormal$, $3$hmiNo$
         Else
           SmartTags("AFEStatus") = "Cannot open file"
         End If  
       End If
     End If
   'Windows / PC based 
   Else
     If SmartTags("aFile_"&SmartTags("AfileChosen")) <> "" Then
       If SmartTags("aIsFolder_"&SmartTags("AfileChosen")) <> "False" Then
         LHmiView_vbsFEReadFilesOfFolder_1(SmartTags("aFile_"&SmartTags("AfileChosen"))&"\")
         LHmiView_vbsFEWriteFilePropertiesToTags_1 1
         SmartTags("Aindex") = 1
       Else  
         fileName = SmartTags("aFile_"&SmartTags("AfileChosen")) 
         Set obj = CreateObject("Wscript.Shell")
         obj.Run fileName
       End If
     Else
       SmartTags("AFEStatus") = "No file or folder chosen"
     End If
   End If

VB script "LHmiView_vbsFEMove_1"
   On Error Resume Next
   
   '-----------------------DEFINE PARAMETERS-------------------------------------------
   'kindOfOperatingSystem: 0 = Windows, 1 = Windows CE
   ' tempFs: Reference on temporary fileSystem Object
   ' fs: Reference on fileSystem Object
   ' f: Reference on file Object
   Dim kindOfOperatingSystem, tempFs, f, fs, file
   
   '--------------------Prove which Operating System is running------------------------
   'Set tempFs = CreateObject("Scripting.FileSystemObject")
   
   'If Err.Number = 0 Then
   '	kindOfOperatingSystem = 0 'Windows / PC based
   'Else
   	kindOfOperatingSystem = 1 'Windows CE / Panel based
   'End If
   
   Set tempFs= Nothing
   Err.Clear
   
   '-------------------------------Move folder/file---------------------------------
   Dim  newpath, singleFile, data
   
   ' Windows CE / Panel based
   If kindOfOperatingSystem Then
     If sender = 1 Then 'button "copy" pressed
   	  If SmartTags("copyusb") = True Then
   		    If SmartTags("IsFolder_"&SmartTags("fileChosen")) = 0 Then
   			      SmartTags("AbufferFile") = SmartTags("File_"&SmartTags("fileChosen"))
   			      SmartTags("AbufferFolder") = SmartTags("Folder")
   			      SmartTags("AbufferCopyCut") = True
   			      SmartTags("AbufferIsFolder") = SmartTags("isFolder_"&SmartTags("fileChosen"))
   			      SmartTags("AFEStatus") = "File " & SmartTags("AbufferFile") & " copied"
   		    Else
   		      	  SmartTags("AFEStatus") = "Cannot copy folder"
   			End If
   	  Else
   		    If SmartTags("AIsFolder_"&SmartTags("AfileChosen")) = 0 Then
   			      SmartTags("AbufferFile") = SmartTags("aFile_"&SmartTags("AfileChosen"))
   			      SmartTags("AbufferFolder") = SmartTags("AFolder")
   			      SmartTags("AbufferCopyCut") = True
   			      SmartTags("AbufferIsFolder") = SmartTags("aisFolder_"&SmartTags("AfileChosen"))
   			      SmartTags("AFEStatus") = "File " & SmartTags("AbufferFile") & " copied"
   		    Else
   		          SmartTags("AFEStatus") = "Cannot copy folder"
   			End If
   	  End If
   	  
     
